// TIA Portal project "XSFW_TIA32801_A0" (V13) (continued)
REGION Network 3: Estado1-->Estado2 (Reposo--> Arranca cinta)
   RUNG wire#powerrail
      Contact( "1s1" )
      Contact( "iSNSpush_atras" )
      wire#w1
      Contact( "iS_automat" )
      wire#w2
      Contact( "iSNS_bs_abajo" )
      Contact( "Marcha" )
      wire#w3
      Contact( "Ya buscó caja" )
      wire#w4
      I_Contact( "Serie de Alarmas" )
      I_Contact( "Cajas acumuladas en salida" )
      Coil( "1c2" )
   END_RUNG
   RUNG wire#powerrail
      Contact( "1s8" )
      Contact( "CERO" )
      I_Contact( "Parada" )
      I_Contact( "Aux acaja acum" )
      I_Contact( "Aux caja trab" )
   END_RUNG wire#w1
   RUNG wire#w1
      Contact( "Modo Manual" )
      I_Contact( "iS_automat" )
      Contact( "fls_Modomanual" )
   END_RUNG wire#w2
   RUNG wire#w3
      Contact( "UNO" )
   END_RUNG wire#w4
   // the same network as SCL:
   "1c2" := (("1s1" AND "iSNSpush_atras") OR ("1s8" AND "CERO" AND NOT "Parada" AND NOT "Aux acaja acum" AND NOT "Aux caja trab")) AND ("iS_automat" OR ("Modo Manual" AND NOT "iS_automat" AND "fls_Modomanual")) AND "iSNS_bs_abajo" AND "Marcha" AND ("Ya buscó caja" OR "UNO") AND NOT "Serie de Alarmas" AND NOT "Cajas acumuladas en salida";
END_REGION

REGION Network 4: Estado2->Estado3 (Arranca Cinta --> Activar retenedores de caja)
   RUNG wire#powerrail
      { S7_Templates := "SrcType := DInt" } GE_Contact(in1 := "Encoder", in2 := 210)
      Contact( "1s2" )
      I_Contact( "Alarmas emergencia y térmicas" )
      I_Contact( "Alarmas cinta" )
      I_Contact( "Serie de Alarmas" )
      Coil( "1c3" )
   END_RUNG
   // the same network as SCL:
   "1c3" := ("Encoder" >= 210) AND "1s2" AND NOT "Alarmas emergencia y térmicas" AND NOT "Alarmas cinta" AND NOT "Serie de Alarmas";
END_REGION

REGION Network 5: Estado3-->Estado4 (Activar retenedores de caja--> Desactivar cinta)
   RUNG wire#powerrail
      Contact( "Punto neutro" )
      Contact( "1s3" )
      I_Contact( "Alarmas emergencia y térmicas" )
      I_Contact( "Alarmas cinta" )
      I_Contact( "Serie de Alarmas" )
      Coil( "1c4" )
   END_RUNG
   RUNG wire#powerrail
      { S7_Templates := "SrcType := DInt" } GE_Contact(in1 := "Encoder", in2 := 238)
      Coil( "Punto neutro" )
   END_RUNG
   // the same network as SCL:
   "1c4" := "Punto neutro" AND "1s3" AND NOT "Alarmas emergencia y térmicas" AND NOT "Alarmas cinta" AND NOT "Serie de Alarmas";
   "Punto neutro" := "Encoder" >= 238;
END_REGION

REGION Network 6: Estado4--> Estado5 (Desactivar cinta--> Activar Pusher y Pinza )
   RUNG wire#powerrail
      Contact( "1s4" )
      Contact( "Auxencol2" )
      I_Contact( "Alarmas"."falla en rele de cadena" )
      I_Contact( "Alarmas emergencia y térmicas" )
      I_Contact( "Alarmas salida y alim de cartones" )
      I_Contact( "Alarmas pusher" )
      I_Contact( "Alarmas brazo de succión" )
      I_Contact( "Serie de Alarmas" )
      Contact( "iSNSpush_atras" )
      Coil( "1c5" )
   END_RUNG
   // the same network as SCL:
   "1c5" := "1s4" AND "Auxencol2" AND NOT "Alarmas"."falla en rele de cadena" AND NOT "Alarmas emergencia y térmicas" AND NOT "Alarmas salida y alim de cartones" AND NOT "Alarmas pusher" AND NOT "Alarmas brazo de succión" AND NOT "Serie de Alarmas" AND "iSNSpush_atras";
END_REGION

REGION Network 7: Estado5-->Estado6 (Activar Pusher y Pinza--> Cilindro Pusher afuera)
   RUNG wire#powerrail
      Contact( "1s5" )
      wire#w1
      Contact( "iSNSalp" )
      I_Contact( "Serie de Alarmas" )
      I_Contact( "Alarmas emergencia y térmicas" )
      I_Contact( "Alarmas pusher" )
      Coil( "1c6" )
   END_RUNG
   RUNG wire#powerrail
      Contact( "CERO" )
      Contact( "1s3" )
      I_Contact( "1c4" )
   END_RUNG wire#w1
   RUNG wire#powerrail
      Contact( "CERO" )
      Contact( "1s4" )
      I_Contact( "1c5" )
   END_RUNG wire#w1
   // the same network as SCL:
   "1c6" := ("1s5" OR ("CERO" AND "1s3" AND NOT "1c4") OR ("CERO" AND "1s4" AND NOT "1c5")) AND "iSNSalp" AND NOT "Serie de Alarmas" AND NOT "Alarmas emergencia y térmicas" AND NOT "Alarmas pusher";
END_REGION

REGION Network 8: Estado6--> Estado7 (Cilindro Pusher afuera--> Desactivar cilindro pusher y pinza )
   RUNG wire#powerrail
      Contact( "1s6" )
      Contact( "iSNSpush_adel" )
      I_Contact( "Serie de Alarmas" )
      I_Contact( "Alarmas emergencia y térmicas" )
      I_Contact( "Alarmas pusher" )
      Coil( "1c7" )
   END_RUNG
   // the same network as SCL:
   "1c7" := "1s6" AND "iSNSpush_adel" AND NOT "Serie de Alarmas" AND NOT "Alarmas emergencia y térmicas" AND NOT "Alarmas pusher";
END_REGION

REGION Network 9: Estado7-->Estado8 (Desactivar cilindro pusher y pinza--> Área libre de Pusher)
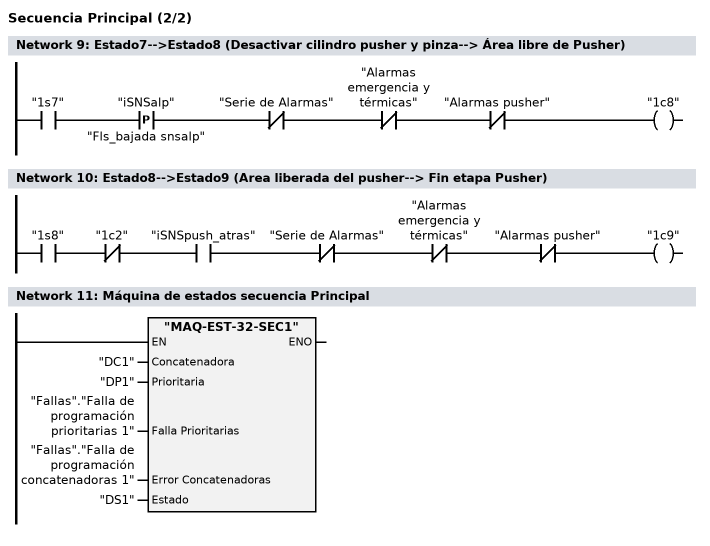
   RUNG wire#powerrail
      Contact( "1s7" )
      P_Contact(operand := "iSNSalp", bit := "Fls_bajada snsalp")
      I_Contact( "Serie de Alarmas" )
      I_Contact( "Alarmas emergencia y térmicas" )
      I_Contact( "Alarmas pusher" )
      Coil( "1c8" )
   END_RUNG
   // the same network as SCL:
   #_w1 := "1s7" AND "iSNSalp" AND NOT "Fls_bajada snsalp";   // rising edge of "iSNSalp"
   "Fls_bajada snsalp" := "iSNSalp";
   "1c8" := #_w1 AND NOT "Serie de Alarmas" AND NOT "Alarmas emergencia y térmicas" AND NOT "Alarmas pusher";
END_REGION

REGION Network 10: Estado8-->Estado9 (Area liberada del pusher--> Fin etapa Pusher)
   RUNG wire#powerrail
      Contact( "1s8" )
      I_Contact( "1c2" )
      Contact( "iSNSpush_atras" )
      I_Contact( "Serie de Alarmas" )
      I_Contact( "Alarmas emergencia y térmicas" )
      I_Contact( "Alarmas pusher" )
      Coil( "1c9" )
   END_RUNG
   // the same network as SCL:
   "1c9" := "1s8" AND NOT "1c2" AND "iSNSpush_atras" AND NOT "Serie de Alarmas" AND NOT "Alarmas emergencia y térmicas" AND NOT "Alarmas pusher";
END_REGION

REGION Network 11: Máquina de estados secuencia Principal
   RUNG wire#powerrail
      "MAQ-EST-32-SEC1"(Concatenadora := "DC1", Prioritaria := "DP1", "Falla Prioritarias" := "Fallas"."Falla de programación prioritarias 1", "Error Concatenadoras" := "Fallas"."Falla de programación concatenadoras 1", Estado := "DS1")
   END_RUNG
   // the same network as SCL:
   "MAQ-EST-32-SEC1"(Concatenadora := "DC1",
                     Prioritaria := "DP1",
                     "Falla Prioritarias" := "Fallas"."Falla de programación prioritarias 1",
                     "Error Concatenadoras" := "Fallas"."Falla de programación concatenadoras 1",
                     Estado := "DS1");
END_REGION
END_FUNCTION

FUNCTION "Condiciones de Marcha y Parada" : Void   // FC7, LAD
TITLE = Condiciones de MARCHA y PARADA (Se la considera una falla prioritaria).
{ S7_Optimized_Access := 'FALSE' }
VERSION : 0.1
// Establece la marcha del proceso según una determinada cantidad de condiciones. En particular para que arranque, se deberá presionar "avería/reposición" . Ya sea que se presione "Parada" o ocurra situaciones de Alarma, se desactivará "Marcha". La diferencia entre ambas es que, para arrancar el sistema luego de una parada, no hace falta presionar nuevamente "avería/reposición". Caso contrario ocurre si quiero arrancar el sistema luego de una Alarma.
BEGIN

REGION Network 1: Condiciones de Marcha
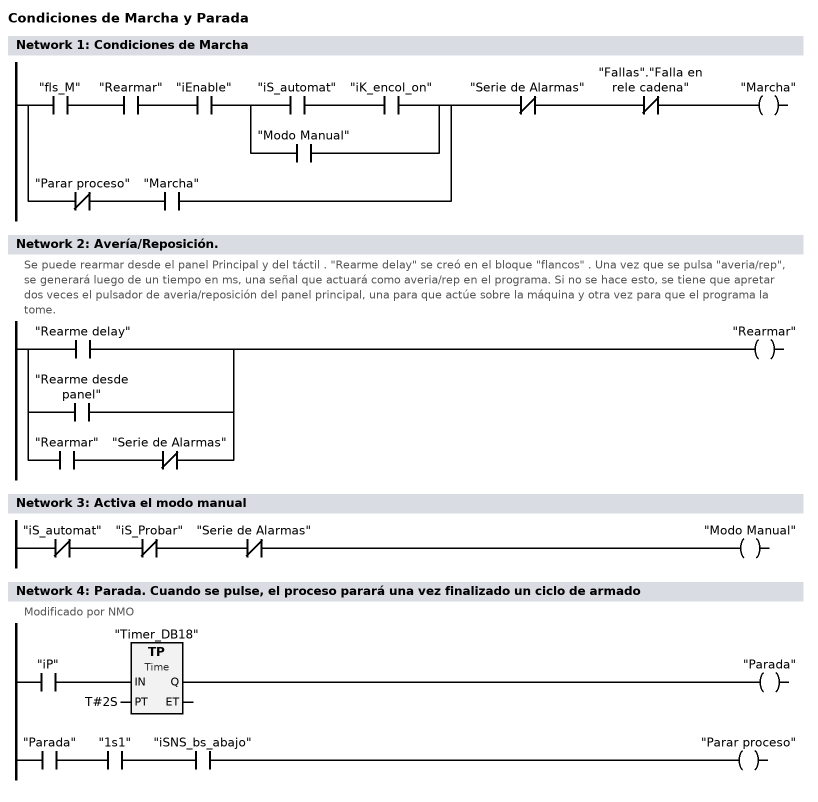
   RUNG wire#powerrail
      Contact( "fls_M" )
      Contact( "Rearmar" )
      Contact( "iEnable" )
      wire#w1
      Contact( "iS_automat" )
      Contact( "iK_encol_on" )
      wire#w2
      I_Contact( "Serie de Alarmas" )
      I_Contact( "Fallas"."Falla en rele cadena" )
      Coil( "Marcha" )
   END_RUNG
   RUNG wire#w1
      Contact( "Modo Manual" )
   END_RUNG wire#w2
   RUNG wire#powerrail
      I_Contact( "Parar proceso" )
      Contact( "Marcha" )
   END_RUNG wire#w2
   // the same network as SCL:
   "Marcha" := (("fls_M" AND "Rearmar" AND "iEnable" AND (("iS_automat" AND "iK_encol_on") OR "Modo Manual")) OR (NOT "Parar proceso" AND "Marcha")) AND NOT "Serie de Alarmas" AND NOT "Fallas"."Falla en rele cadena";
END_REGION

REGION Network 2: Avería/Reposición.
   // Se puede rearmar desde el panel Principal y del táctil . "Rearme delay" se creó en el bloque "flancos" . Una vez que se pulsa "averia/rep", se generará luego de un tiempo en ms, una señal que actuará como averia/rep en el programa. Si no se hace esto, se tiene que apretar dos veces el pulsador de averia/reposición del panel principal, una para que actúe sobre la máquina y otra vez para que el programa la tome.
   RUNG wire#powerrail
      Contact( "Rearme delay" )
      wire#w1
      Coil( "Rearmar" )
   END_RUNG
   RUNG wire#powerrail
      Contact( "Rearme desde panel" )
   END_RUNG wire#w1
   RUNG wire#powerrail
      Contact( "Rearmar" )
      I_Contact( "Serie de Alarmas" )
   END_RUNG wire#w1
   // the same network as SCL:
   "Rearmar" := "Rearme delay" OR "Rearme desde panel" OR ("Rearmar" AND NOT "Serie de Alarmas");
END_REGION

REGION Network 3: Activa el modo manual
   RUNG wire#powerrail
      I_Contact( "iS_automat" )
      I_Contact( "iS_Probar" )
      I_Contact( "Serie de Alarmas" )
      Coil( "Modo Manual" )
   END_RUNG
   // the same network as SCL:
   "Modo Manual" := NOT "iS_automat" AND NOT "iS_Probar" AND NOT "Serie de Alarmas";
END_REGION

REGION Network 4: Parada. Cuando se pulse, el proceso parará una vez finalizado un ciclo de armado
   // Modificado por NMO
   "Timer_DB18".TP(IN := "iP", PT := T#2S);
   "Parada" := "Timer_DB18".Q;
   "Parar proceso" := "Parada" AND "1s1" AND "iSNS_bs_abajo";
END_REGION
END_FUNCTION

FUNCTION "Contador rápido y encoder" : Void   // FC8, LAD
TITLE = Lleva la cuenta de los pulsos del ENCODER.
{ S7_Optimized_Access := 'FALSE' }
VERSION : 0.1
   VAR_TEMP   // added for the SCL form of the ladder/FBD networks
      _w1 : Bool;
   END_VAR
BEGIN

REGION Network 1: Reset del HSC para poner en cero el encóder.
   // En HSC va 258, es la ID de Hardware
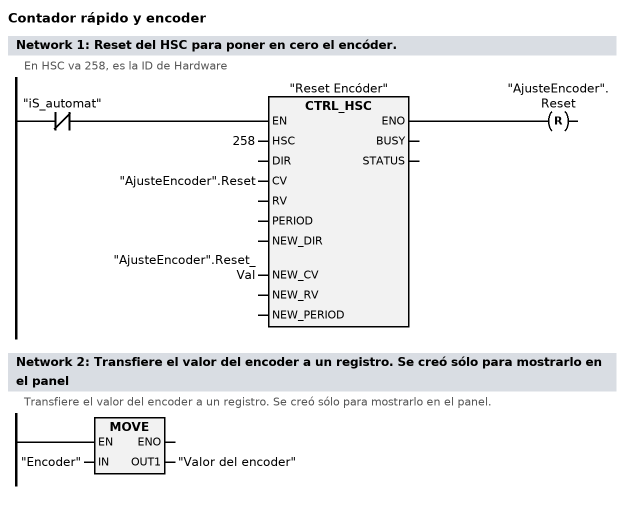
   // ENO of a box is taken as its EN; it also drops when the box reports an error
   #_w1 := NOT "iS_automat";
   IF #_w1 THEN
       "Reset Encóder"(HSC := 258, CV := "AjusteEncoder".Reset, NEW_CV := "AjusteEncoder".Reset_Val);   // CTRL_HSC
       "AjusteEncoder".Reset := FALSE;
   END_IF;
END_REGION

REGION Network 2: Transfiere el valor del encoder a un registro. Se creó sólo para mostrarlo en el panel
   // Transfiere el valor del encoder a un registro. Se creó sólo para mostrarlo en el panel.
   RUNG wire#powerrail
      { S7_GenerateENO := "TRUE" } Move(in := "Encoder", out1 => "Valor del encoder")
   END_RUNG
   // the same network as SCL:
   "Valor del encoder" := "Encoder";
END_REGION
END_FUNCTION

FUNCTION "cajas armadas hasta el momento" : Void   // FC9, LAD
{ S7_Optimized_Access := 'FALSE' }
VERSION : 0.1
BEGIN

REGION Network 1: Contabiliza la cantidad de cajas armadas.
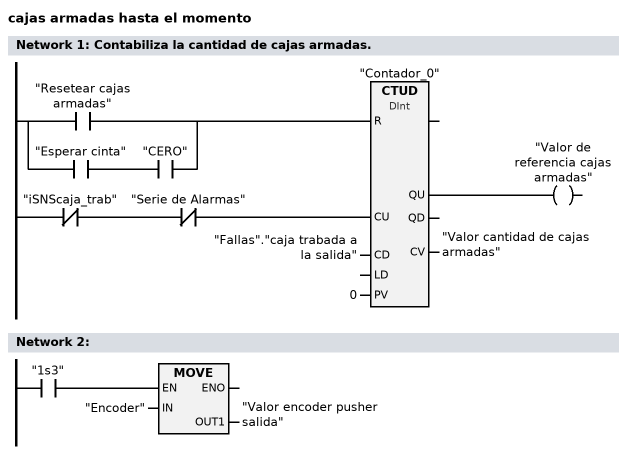
   "Contador_0".CTUD(cu := NOT "iSNScaja_trab" AND NOT "Serie de Alarmas",
                     r := "Resetear cajas armadas" OR ("Esperar cinta" AND "CERO"),
                     cd := "Fallas"."caja trabada a la salida",
                     pv := 0,
                     cv => "Valor cantidad de cajas armadas");
   "Valor de referencia cajas armadas" := "Contador_0".qu;
END_REGION

REGION Network 2
   RUNG wire#powerrail
      Contact( "1s3" )
      { S7_GenerateENO := "TRUE" } Move(in := "Encoder", out1 => "Valor encoder pusher salida")
   END_RUNG
   // the same network as SCL:
   IF "1s3" THEN "Valor encoder pusher salida" := "Encoder"; END_IF;
END_REGION
END_FUNCTION

FUNCTION "Luces de marcha y parada" : Void   // FC10, LAD
{ S7_Optimized_Access := 'FALSE' }
VERSION : 0.1
BEGIN

REGION Network 1: Luz de Marcha
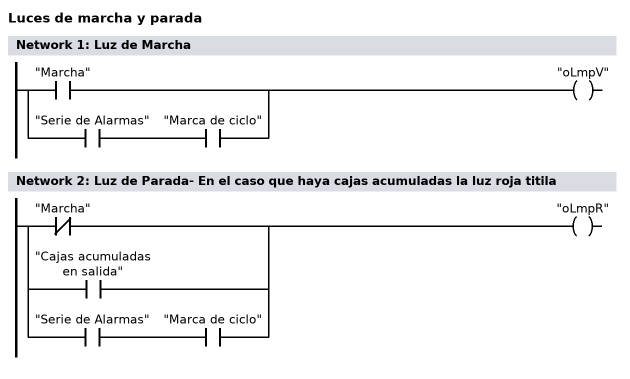
   RUNG wire#powerrail
      Contact( "Marcha" )
      wire#w1
      Coil( "oLmpV" )
   END_RUNG
   RUNG wire#powerrail
      Contact( "Serie de Alarmas" )
      Contact( "Marca de ciclo" )
   END_RUNG wire#w1
   // the same network as SCL:
   "oLmpV" := "Marcha" OR ("Serie de Alarmas" AND "Marca de ciclo");
END_REGION

REGION Network 2: Luz de Parada- En el caso que haya cajas acumuladas la luz roja titila
   RUNG wire#powerrail
      I_Contact( "Marcha" )
      wire#w1
      Coil( "oLmpR" )
   END_RUNG
   RUNG wire#powerrail
      Contact( "Cajas acumuladas en salida" )
   END_RUNG wire#w1
   RUNG wire#powerrail
      Contact( "Serie de Alarmas" )
      Contact( "Marca de ciclo" )
   END_RUNG wire#w1
   // the same network as SCL:
   "oLmpR" := NOT "Marcha" OR "Cajas acumuladas en salida" OR ("Serie de Alarmas" AND "Marca de ciclo");
END_REGION
END_FUNCTION

FUNCTION "flancos" : Void   // FC12, LAD
{ S7_Optimized_Access := 'FALSE' }
VERSION : 0.1
   VAR_TEMP   // added for the SCL form of the ladder/FBD networks
      _w1 : Bool;
   END_VAR
BEGIN

REGION Network 1: avería/ reposición
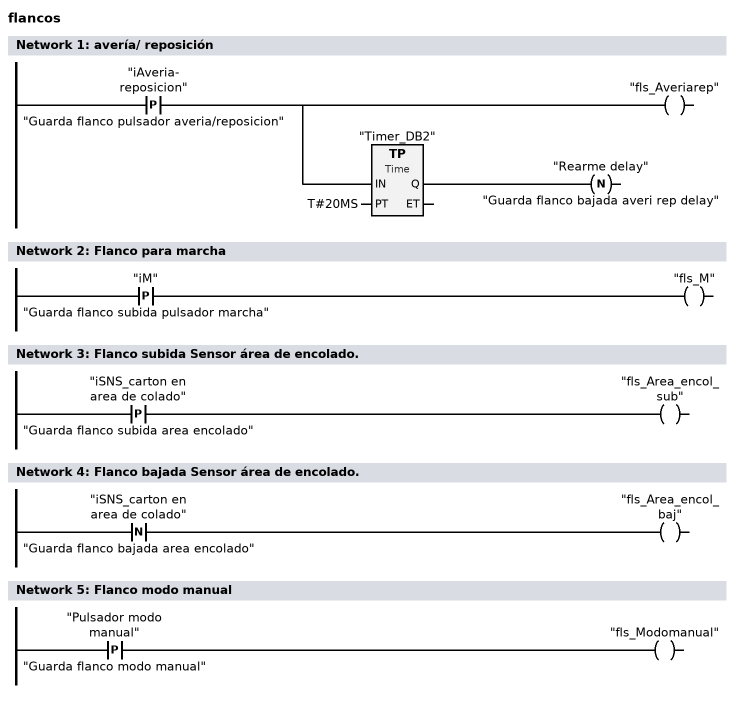
   #_w1 := "iAveria-reposicion" AND NOT "Guarda flanco pulsador averia/reposicion";   // rising edge of "iAveria-reposicion"
   "Guarda flanco pulsador averia/reposicion" := "iAveria-reposicion";
   "fls_Averiarep" := #_w1;
   "Timer_DB2".TP(in := #_w1, pt := T#20MS);
   "Rearme delay" := NOT "Timer_DB2".q AND "Guarda flanco bajada averi rep delay";   // falling edge
   "Guarda flanco bajada averi rep delay" := "Timer_DB2".q;
END_REGION

REGION Network 2: Flanco para marcha
   RUNG wire#powerrail
      P_Contact(operand := "iM", bit := "Guarda flanco subida pulsador marcha")
      Coil( "fls_M" )
   END_RUNG
   // the same network as SCL:
   #_w1 := "iM" AND NOT "Guarda flanco subida pulsador marcha";   // rising edge of "iM"
   "Guarda flanco subida pulsador marcha" := "iM";
   "fls_M" := #_w1;
END_REGION

REGION Network 3: Flanco subida Sensor área de encolado.
   RUNG wire#powerrail
      P_Contact(operand := "iSNS_carton en area de colado", bit := "Guarda flanco subida area encolado")
      Coil( "fls_Area_encol_sub" )
   END_RUNG
   // the same network as SCL:
   #_w1 := "iSNS_carton en area de colado" AND NOT "Guarda flanco subida area encolado";   // rising edge of "iSNS_carton en area de colado"
   "Guarda flanco subida area encolado" := "iSNS_carton en area de colado";
   "fls_Area_encol_sub" := #_w1;
END_REGION

REGION Network 4: Flanco bajada Sensor área de encolado.
   RUNG wire#powerrail
      N_Contact(operand := "iSNS_carton en area de colado", bit := "Guarda flanco bajada area encolado")
      Coil( "fls_Area_encol_baj" )
   END_RUNG
   // the same network as SCL:
   #_w1 := NOT "iSNS_carton en area de colado" AND "Guarda flanco bajada area encolado";   // falling edge of "iSNS_carton en area de colado"
   "Guarda flanco bajada area encolado" := "iSNS_carton en area de colado";
   "fls_Area_encol_baj" := #_w1;
END_REGION

REGION Network 5: Flanco modo manual
   RUNG wire#powerrail
      P_Contact(operand := "Pulsador modo manual", bit := "Guarda flanco modo manual")
      Coil( "fls_Modomanual" )
   END_RUNG
   // the same network as SCL:
   #_w1 := "Pulsador modo manual" AND NOT "Guarda flanco modo manual";   // rising edge of "Pulsador modo manual"
   "Guarda flanco modo manual" := "Pulsador modo manual";
   "fls_Modomanual" := #_w1;
END_REGION
END_FUNCTION

FUNCTION "MODO PROBAR (MP)" : Void   // FC13, LAD
{ S7_Optimized_Access := 'FALSE' }
VERSION : 0.1
   VAR_TEMP   // added for the SCL form of the ladder/FBD networks
      _w1 : Bool;
   END_VAR
BEGIN

REGION Network 1: Modo Probar. En este caso se desactivan las alarmas excepto la de emergencia y térmicas.
   // Si no está en automático, y no hay alarmas, se activa el modo PROBAR. Con esto se activa la bomba de vacío.
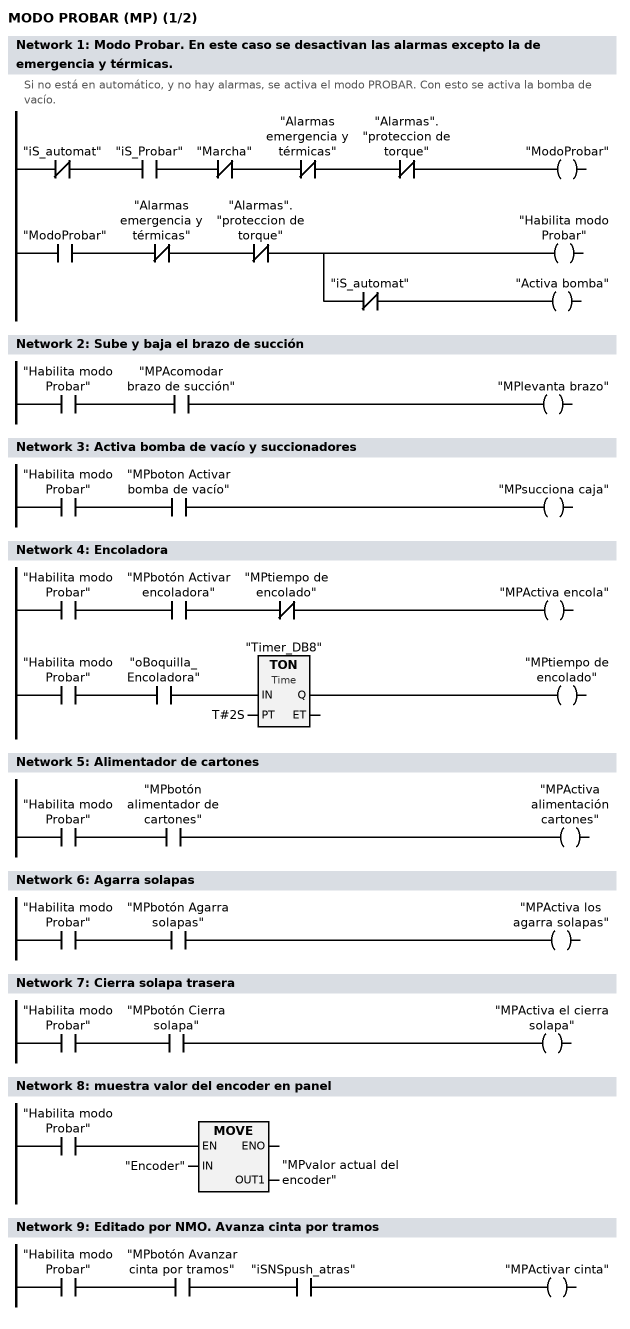
   RUNG wire#powerrail
      I_Contact( "iS_automat" )
      Contact( "iS_Probar" )
      I_Contact( "Marcha" )
      I_Contact( "Alarmas emergencia y térmicas" )
      I_Contact( "Alarmas"."proteccion de torque" )
      Coil( "ModoProbar" )
   END_RUNG
   RUNG wire#powerrail
      Contact( "ModoProbar" )
      I_Contact( "Alarmas emergencia y térmicas" )
      I_Contact( "Alarmas"."proteccion de torque" )
      wire#w1
      Coil( "Habilita modo Probar" )
   END_RUNG
   RUNG wire#w1
      I_Contact( "iS_automat" )
      Coil( "Activa bomba" )
   END_RUNG
   // the same network as SCL:
   "ModoProbar" := NOT "iS_automat" AND "iS_Probar" AND NOT "Marcha" AND NOT "Alarmas emergencia y térmicas" AND NOT "Alarmas"."proteccion de torque";
   "Habilita modo Probar" := "ModoProbar" AND NOT "Alarmas emergencia y térmicas" AND NOT "Alarmas"."proteccion de torque";
   "Activa bomba" := "Habilita modo Probar" AND NOT "iS_automat";
END_REGION

REGION Network 2: Sube y baja el brazo de succión
   RUNG wire#powerrail
      Contact( "Habilita modo Probar" )
      Contact( "MPAcomodar brazo de succión" )
      Coil( "MPlevanta brazo" )
   END_RUNG
   // the same network as SCL:
   "MPlevanta brazo" := "Habilita modo Probar" AND "MPAcomodar brazo de succión";
END_REGION

REGION Network 3: Activa bomba de vacío y succionadores
   RUNG wire#powerrail
      Contact( "Habilita modo Probar" )
      Contact( "MPboton Activar bomba de vacío" )
      Coil( "MPsucciona caja" )
   END_RUNG
   // the same network as SCL:
   "MPsucciona caja" := "Habilita modo Probar" AND "MPboton Activar bomba de vacío";
END_REGION

REGION Network 4: Encoladora
   "MPActiva encola" := "Habilita modo Probar" AND "MPbotón Activar encoladora" AND NOT "MPtiempo de encolado";
   "Timer_DB8".TON(IN := "Habilita modo Probar" AND "oBoquilla_Encoladora", PT := T#2S);
   "MPtiempo de encolado" := "Timer_DB8".Q;
END_REGION

REGION Network 5: Alimentador de cartones
   RUNG wire#powerrail
      Contact( "Habilita modo Probar" )
      Contact( "MPbotón alimentador de cartones" )
      Coil( "MPActiva alimentación cartones" )
   END_RUNG
   // the same network as SCL:
   "MPActiva alimentación cartones" := "Habilita modo Probar" AND "MPbotón alimentador de cartones";
END_REGION

REGION Network 6: Agarra solapas
   RUNG wire#powerrail
      Contact( "Habilita modo Probar" )
      Contact( "MPbotón Agarra solapas" )
      Coil( "MPActiva los agarra solapas" )
   END_RUNG
   // the same network as SCL:
   "MPActiva los agarra solapas" := "Habilita modo Probar" AND "MPbotón Agarra solapas";
END_REGION

REGION Network 7: Cierra solapa trasera
   RUNG wire#powerrail
      Contact( "Habilita modo Probar" )
      Contact( "MPbotón Cierra solapa" )
      Coil( "MPActiva el cierra solapa" )
   END_RUNG
   // the same network as SCL:
   "MPActiva el cierra solapa" := "Habilita modo Probar" AND "MPbotón Cierra solapa";
END_REGION

REGION Network 8: muestra valor del encoder en panel
   RUNG wire#powerrail
      Contact( "Habilita modo Probar" )
      { S7_GenerateENO := "TRUE" } Move(in := "Encoder", out1 => "MPvalor actual del encoder")
   END_RUNG
   // the same network as SCL:
   IF "Habilita modo Probar" THEN "MPvalor actual del encoder" := "Encoder"; END_IF;
END_REGION

REGION Network 9: Editado por NMO. Avanza cinta por tramos
   RUNG wire#powerrail
      Contact( "Habilita modo Probar" )
      Contact( "MPbotón Avanzar cinta por tramos" )
      Contact( "iSNSpush_atras" )
      Coil( "MPActivar cinta" )
   END_RUNG
   // the same network as SCL:
   "MPActivar cinta" := "Habilita modo Probar" AND "MPbotón Avanzar cinta por tramos" AND "iSNSpush_atras";
END_REGION

REGION Network 10: Editado por NMO. Desactivar marca "MPbotón avanzar cinta por tramos".
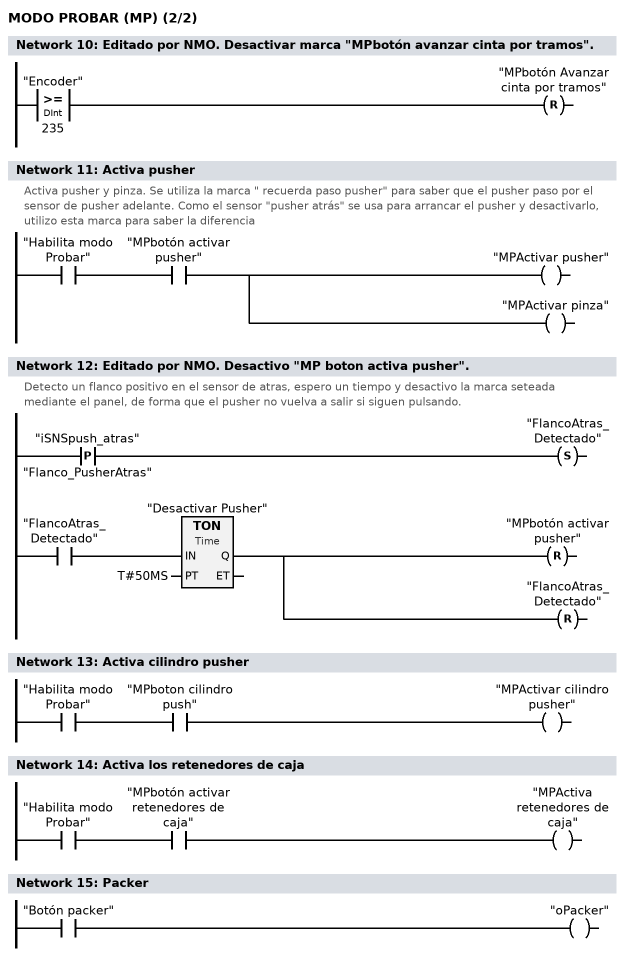
   RUNG wire#powerrail
      { S7_Templates := "SrcType := DInt" } GE_Contact(in1 := "Encoder", in2 := 235)
      R_Coil( "MPbotón Avanzar cinta por tramos" )
   END_RUNG
   // the same network as SCL:
   IF "Encoder" >= 235 THEN "MPbotón Avanzar cinta por tramos" := FALSE; END_IF;
END_REGION

REGION Network 11: Activa pusher
   // Activa pusher y pinza. Se utiliza la marca " recuerda paso pusher" para saber que el pusher paso por el sensor de pusher adelante. Como el sensor "pusher atrás" se usa para arrancar el pusher y desactivarlo, utilizo esta marca para saber la diferencia
   RUNG wire#powerrail
      Contact( "Habilita modo Probar" )
      Contact( "MPbotón activar pusher" )
      wire#w1
      Coil( "MPActivar pusher" )
   END_RUNG
   RUNG wire#w1
      Coil( "MPActivar pinza" )
   END_RUNG
   // the same network as SCL:
   "MPActivar pusher" := "Habilita modo Probar" AND "MPbotón activar pusher";
   "MPActivar pinza" := "MPActivar pusher";
END_REGION

REGION Network 12: Editado por NMO. Desactivo "MP boton activa pusher".
   // Detecto un flanco positivo en el sensor de atras, espero un tiempo y desactivo la marca seteada mediante el panel, de forma que el pusher no vuelva a salir si siguen pulsando.
   #_w1 := "iSNSpush_atras" AND NOT "Flanco_PusherAtras";   // rising edge of "iSNSpush_atras"
   "Flanco_PusherAtras" := "iSNSpush_atras";
   IF #_w1 THEN "FlancoAtras_Detectado" := TRUE; END_IF;
   "Desactivar Pusher".TON(IN := "FlancoAtras_Detectado", PT := T#50MS);
   IF "Desactivar Pusher".Q THEN
       "MPbotón activar pusher" := FALSE;
       "FlancoAtras_Detectado" := FALSE;
   END_IF;
END_REGION

REGION Network 13: Activa cilindro pusher
   RUNG wire#powerrail
      Contact( "Habilita modo Probar" )
      Contact( "MPboton cilindro push" )
      Coil( "MPActivar cilindro pusher" )
   END_RUNG
   // the same network as SCL:
   "MPActivar cilindro pusher" := "Habilita modo Probar" AND "MPboton cilindro push";
END_REGION

REGION Network 14: Activa los retenedores de caja
   RUNG wire#powerrail
      Contact( "Habilita modo Probar" )
      Contact( "MPbotón activar retenedores de caja" )
      Coil( "MPActiva retenedores de caja" )
   END_RUNG
   // the same network as SCL:
   "MPActiva retenedores de caja" := "Habilita modo Probar" AND "MPbotón activar retenedores de caja";
END_REGION

REGION Network 15: Packer
   RUNG wire#powerrail
      Contact( "Botón packer" )
      Coil( "oPacker" )
   END_RUNG
   // the same network as SCL:
   "oPacker" := "Botón packer";
END_REGION
END_FUNCTION

FUNCTION "Tratamiento de Fallas" : Void   // FC16, LAD
TITLE = Tratamiento de fallas.
{ S7_Optimized_Access := 'FALSE' }
VERSION : 0.1
   VAR_TEMP   // added for the SCL form of the ladder/FBD networks
      _w1 : Bool;
   END_VAR
BEGIN

REGION Network 1: Falla en térmicas.
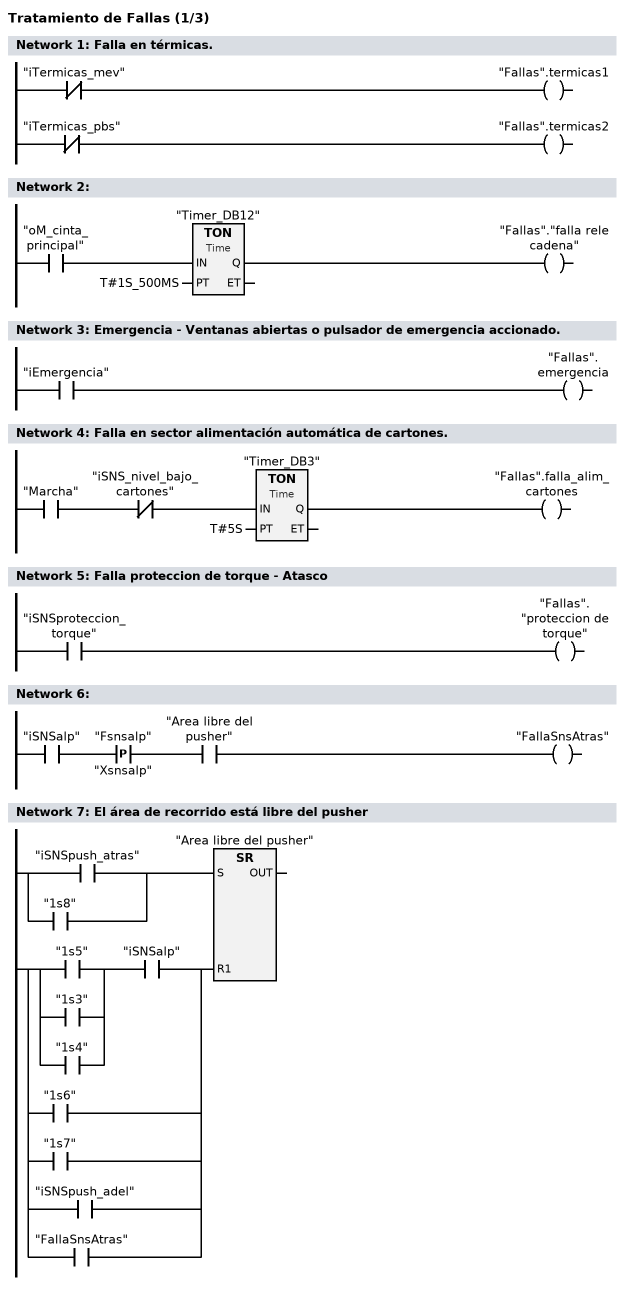
   RUNG wire#powerrail
      I_Contact( "iTermicas_mev" )
      Coil( "Fallas".termicas1 )
   END_RUNG
   RUNG wire#powerrail
      I_Contact( "iTermicas_pbs" )
      Coil( "Fallas".termicas2 )
   END_RUNG
   // the same network as SCL:
   "Fallas".termicas1 := NOT "iTermicas_mev";
   "Fallas".termicas2 := NOT "iTermicas_pbs";
END_REGION

REGION Network 2
   "Timer_DB12".TON(IN := "oM_cinta_principal", PT := T#1S_500MS);
   "Fallas"."falla rele cadena" := "Timer_DB12".Q;
END_REGION

REGION Network 3: Emergencia - Ventanas abiertas o pulsador de emergencia accionado.
   RUNG wire#powerrail
      Contact( "iEmergencia" )
      Coil( "Fallas".emergencia )
   END_RUNG
   // the same network as SCL:
   "Fallas".emergencia := "iEmergencia";
END_REGION

REGION Network 4: Falla en sector alimentación automática de cartones.
   "Timer_DB3".TON(IN := "Marcha" AND NOT "iSNS_nivel_bajo_cartones", PT := T#5S);
   "Fallas".falla_alim_cartones := "Timer_DB3".Q;
END_REGION

REGION Network 5: Falla proteccion de torque - Atasco
   RUNG wire#powerrail
      Contact( "iSNSproteccion_torque" )
      Coil( "Fallas"."proteccion de torque" )
   END_RUNG
   // the same network as SCL:
   "Fallas"."proteccion de torque" := "iSNSproteccion_torque";
END_REGION

REGION Network 6
   RUNG wire#powerrail
      Contact( "iSNSalp" )
      P_Contact(operand := "Fsnsalp", bit := "Xsnsalp")
      Contact( "Area libre del pusher" )
      Coil( "FallaSnsAtras" )
   END_RUNG
   // the same network as SCL:
   #_w1 := "iSNSalp" AND "Fsnsalp" AND NOT "Xsnsalp";   // rising edge of "Fsnsalp"
   "Xsnsalp" := "Fsnsalp";
   "FallaSnsAtras" := #_w1 AND "Area libre del pusher";
END_REGION

REGION Network 7: El área de recorrido está libre del pusher
   RUNG wire#powerrail
      Contact( "iSNSpush_atras" )
      wire#w1
      S_SR(operand := "Area libre del pusher", r1 := wire#w3)
   END_RUNG
   RUNG wire#powerrail
      Contact( "1s8" )
   END_RUNG wire#w1
   RUNG wire#powerrail
      Contact( "1s5" )
      wire#w2
      Contact( "iSNSalp" )
   END_RUNG wire#w3
   RUNG wire#powerrail
      Contact( "1s3" )
   END_RUNG wire#w2
   RUNG wire#powerrail
      Contact( "1s4" )
   END_RUNG wire#w2
   RUNG wire#powerrail
      Contact( "1s6" )
   END_RUNG wire#w3
   RUNG wire#powerrail
      Contact( "1s7" )
   END_RUNG wire#w3
   RUNG wire#powerrail
      Contact( "iSNSpush_adel" )
   END_RUNG wire#w3
   RUNG wire#powerrail
      Contact( "FallaSnsAtras" )
   END_RUNG wire#w3
   // the same network as SCL:
   IF "iSNSpush_atras" OR "1s8" THEN
       "Area libre del pusher" := TRUE;   // SR flip-flop
   END_IF;
   IF (("1s5" OR "1s3" OR "1s4") AND "iSNSalp") OR "1s6" OR "1s7" OR "iSNSpush_adel" OR "FallaSnsAtras" THEN
       "Area libre del pusher" := FALSE;
   END_IF;
END_REGION

REGION Network 8: Incongruencia en sensores del pusher.
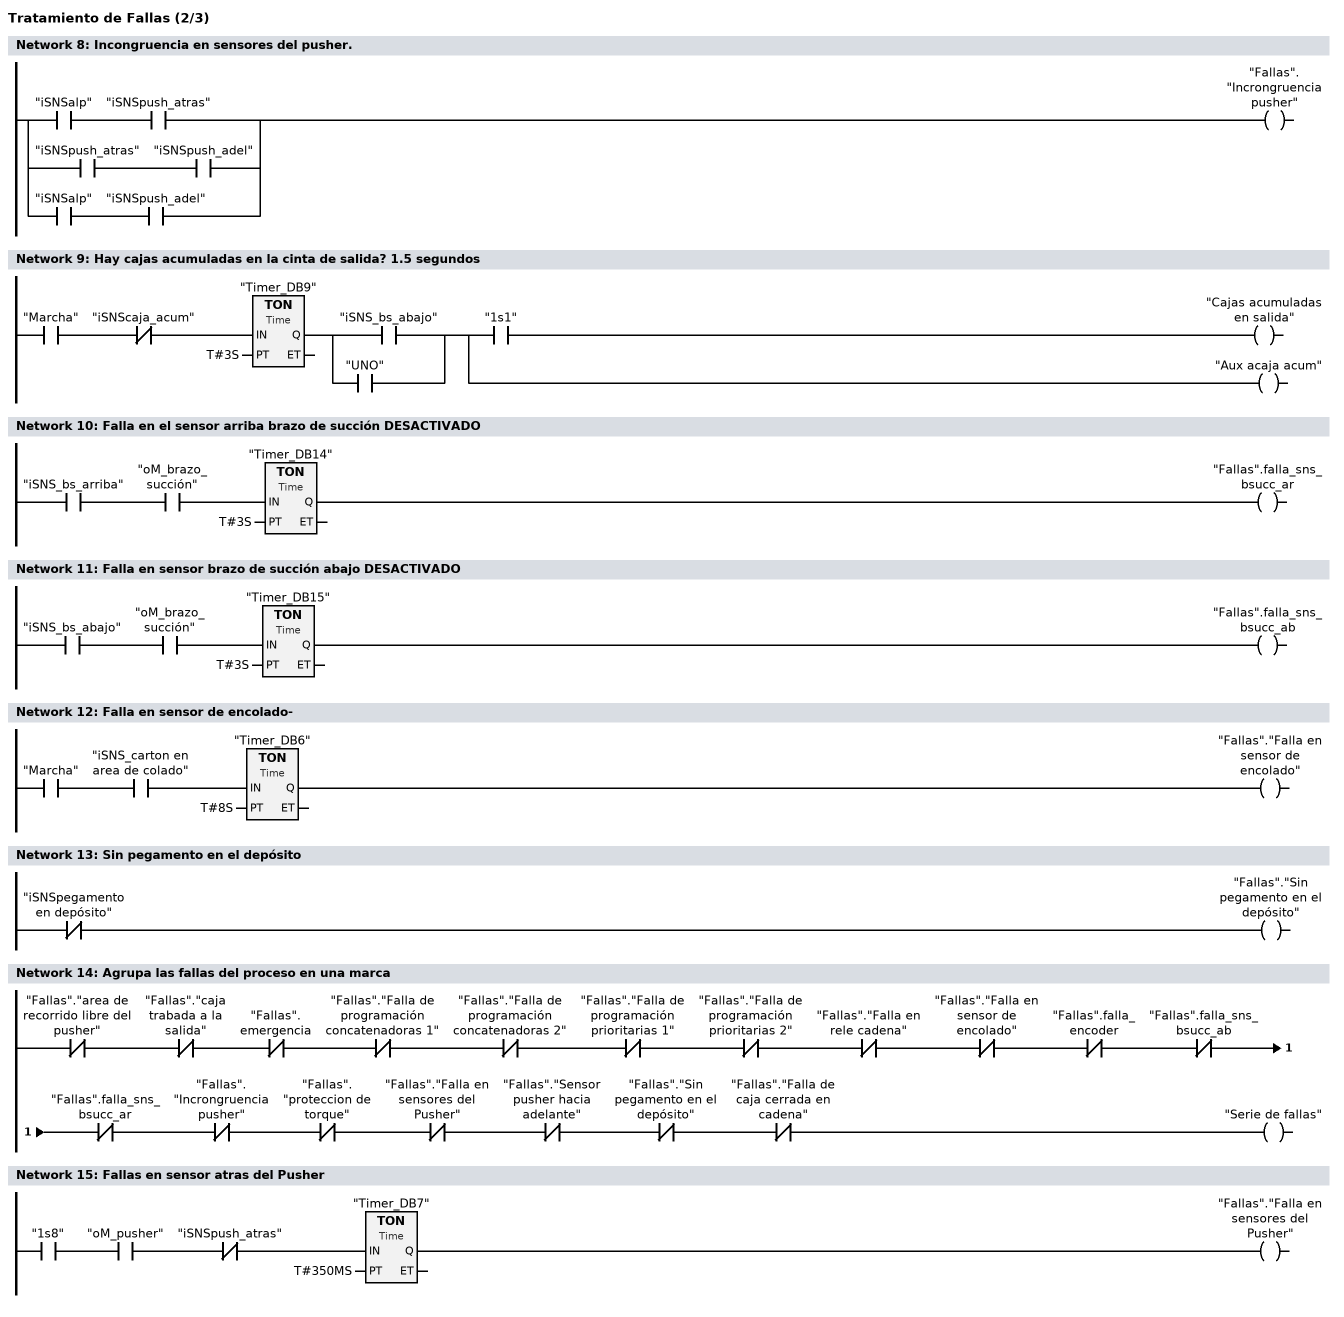
   RUNG wire#powerrail
      Contact( "iSNSalp" )
      Contact( "iSNSpush_atras" )
      wire#w1
      Coil( "Fallas"."Incrongruencia pusher" )
   END_RUNG
   RUNG wire#powerrail
      Contact( "iSNSpush_atras" )
      Contact( "iSNSpush_adel" )
   END_RUNG wire#w1
   RUNG wire#powerrail
      Contact( "iSNSalp" )
      Contact( "iSNSpush_adel" )
   END_RUNG wire#w1
   // the same network as SCL:
   "Fallas"."Incrongruencia pusher" := ("iSNSalp" AND "iSNSpush_atras") OR ("iSNSpush_atras" AND "iSNSpush_adel") OR ("iSNSalp" AND "iSNSpush_adel");
END_REGION

REGION Network 9: Hay cajas acumuladas en la cinta de salida? 1.5 segundos
   "Timer_DB9".TON(in := "Marcha" AND NOT "iSNScaja_acum", pt := T#3S);
   #_w1 := "Timer_DB9".q AND ("iSNS_bs_abajo" OR "UNO");
   "Cajas acumuladas en salida" := #_w1 AND "1s1";
   "Aux acaja acum" := #_w1;
END_REGION

REGION Network 10: Falla en el sensor arriba brazo de succión DESACTIVADO
   "Timer_DB14".TON(IN := "iSNS_bs_arriba" AND "oM_brazo_succión", PT := T#3S);
   "Fallas".falla_sns_bsucc_ar := "Timer_DB14".Q;
END_REGION

REGION Network 11: Falla en sensor brazo de succión abajo DESACTIVADO
   "Timer_DB15".TON(IN := "iSNS_bs_abajo" AND "oM_brazo_succión", PT := T#3S);
   "Fallas".falla_sns_bsucc_ab := "Timer_DB15".Q;
END_REGION

REGION Network 12: Falla en sensor de encolado-
   "Timer_DB6".TON(IN := "Marcha" AND "iSNS_carton en area de colado", PT := T#8S);
   "Fallas"."Falla en sensor de encolado" := "Timer_DB6".Q;
END_REGION

REGION Network 13: Sin pegamento en el depósito
   RUNG wire#powerrail
      I_Contact( "iSNSpegamento en depósito" )
      Coil( "Fallas"."Sin pegamento en el depósito" )
   END_RUNG
   // the same network as SCL:
   "Fallas"."Sin pegamento en el depósito" := NOT "iSNSpegamento en depósito";
END_REGION

REGION Network 14: Agrupa las fallas del proceso en una marca
   RUNG wire#powerrail
      I_Contact( "Fallas"."area de recorrido libre del pusher" )
      I_Contact( "Fallas"."caja trabada a la salida" )
      I_Contact( "Fallas".emergencia )
      I_Contact( "Fallas"."Falla de programación concatenadoras 1" )
      I_Contact( "Fallas"."Falla de programación concatenadoras 2" )
      I_Contact( "Fallas"."Falla de programación prioritarias 1" )
      I_Contact( "Fallas"."Falla de programación prioritarias 2" )
      I_Contact( "Fallas"."Falla en rele cadena" )
      I_Contact( "Fallas"."Falla en sensor de encolado" )
      I_Contact( "Fallas".falla_encoder )
      I_Contact( "Fallas".falla_sns_bsucc_ab )
      I_Contact( "Fallas".falla_sns_bsucc_ar )
      I_Contact( "Fallas"."Incrongruencia pusher" )
      I_Contact( "Fallas"."proteccion de torque" )
      I_Contact( "Fallas"."Falla en sensores del Pusher" )
      I_Contact( "Fallas"."Sensor pusher hacia adelante" )
      I_Contact( "Fallas"."Sin pegamento en el depósito" )
      I_Contact( "Fallas"."Falla de caja cerrada en cadena" )
      Coil( "Serie de fallas" )
   END_RUNG
   // the same network as SCL:
   "Serie de fallas" := NOT "Fallas"."area de recorrido libre del pusher" AND NOT "Fallas"."caja trabada a la salida" AND NOT "Fallas".emergencia AND NOT "Fallas"."Falla de programación concatenadoras 1" AND NOT "Fallas"."Falla de programación concatenadoras 2" AND NOT "Fallas"."Falla de programación prioritarias 1" AND NOT "Fallas"."Falla de programación prioritarias 2" AND NOT "Fallas"."Falla en rele cadena" AND NOT "Fallas"."Falla en sensor de encolado" AND NOT "Fallas".falla_encoder AND NOT "Fallas".falla_sns_bsucc_ab AND NOT "Fallas".falla_sns_bsucc_ar AND NOT "Fallas"."Incrongruencia pusher" AND NOT "Fallas"."proteccion de torque" AND NOT "Fallas"."Falla en sensores del Pusher" AND NOT "Fallas"."Sensor pusher hacia adelante" AND NOT "Fallas"."Sin pegamento en el depósito" AND NOT "Fallas"."Falla de caja cerrada en cadena";
END_REGION

REGION Network 15: Fallas en sensor atras del Pusher
   "Timer_DB7".TON(IN := "1s8" AND "oM_pusher" AND NOT "iSNSpush_atras", PT := T#350MS);
   "Fallas"."Falla en sensores del Pusher" := "Timer_DB7".Q;
END_REGION

REGION Network 16: Fallas en sensor adelante del Pusher
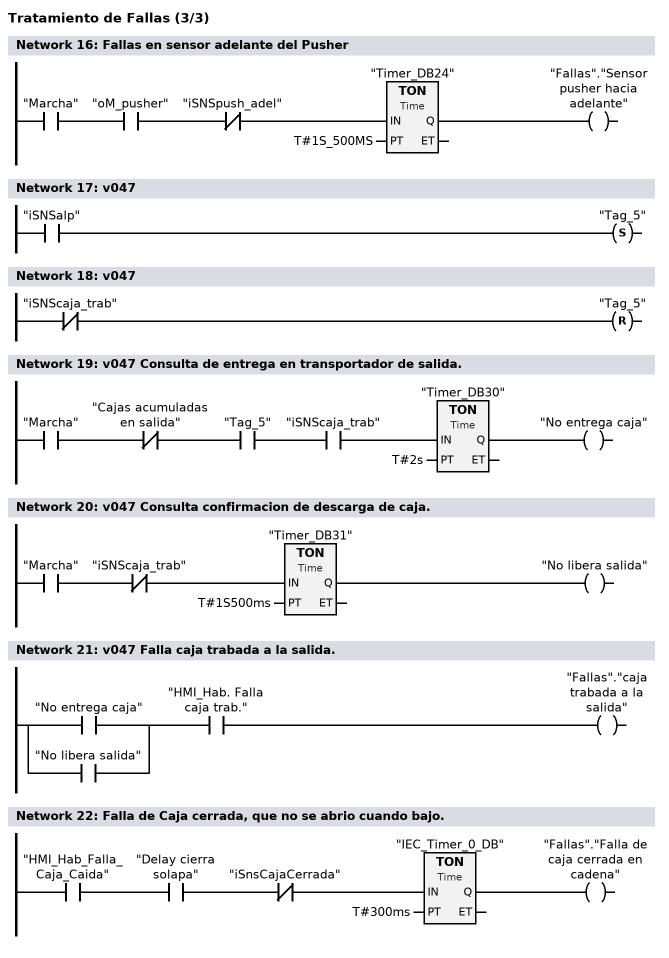
   "Timer_DB24".TON(IN := "Marcha" AND "oM_pusher" AND NOT "iSNSpush_adel", PT := T#1S_500MS);
   "Fallas"."Sensor pusher hacia adelante" := "Timer_DB24".Q;
END_REGION

REGION Network 17: v047
   RUNG wire#powerrail
      Contact( "iSNSalp" )
      S_Coil( "Tag_5" )
   END_RUNG
   // the same network as SCL:
   IF "iSNSalp" THEN "Tag_5" := TRUE; END_IF;
END_REGION

REGION Network 18: v047
   RUNG wire#powerrail
      I_Contact( "iSNScaja_trab" )
      R_Coil( "Tag_5" )
   END_RUNG
   // the same network as SCL:
   IF NOT "iSNScaja_trab" THEN "Tag_5" := FALSE; END_IF;
END_REGION

REGION Network 19: v047 Consulta de entrega en transportador de salida.
   "Timer_DB30".TON(IN := "Marcha" AND NOT "Cajas acumuladas en salida" AND "Tag_5" AND "iSNScaja_trab",
                    PT := T#2s);
   "No entrega caja" := "Timer_DB30".Q;
END_REGION

REGION Network 20: v047 Consulta confirmacion de descarga de caja.
   "Timer_DB31".TON(IN := "Marcha" AND NOT "iSNScaja_trab", PT := T#1S500ms);
   "No libera salida" := "Timer_DB31".Q;
END_REGION

REGION Network 21: v047 Falla caja trabada a la salida.
   RUNG wire#powerrail
      Contact( "No entrega caja" )
      wire#w1
      Contact( "HMI_Hab. Falla caja trab." )
      Coil( "Fallas"."caja trabada a la salida" )
   END_RUNG
   RUNG wire#powerrail
      Contact( "No libera salida" )
   END_RUNG wire#w1
   // the same network as SCL:
   "Fallas"."caja trabada a la salida" := ("No entrega caja" OR "No libera salida") AND "HMI_Hab. Falla caja trab.";
END_REGION

REGION Network 22: Falla de Caja cerrada, que no se abrio cuando bajo.
   "IEC_Timer_0_DB".TON(IN := "HMI_Hab_Falla_Caja_Caida" AND "Delay cierra solapa" AND NOT "iSnsCajaCerrada",
                        PT := T#300ms);
   "Fallas"."Falla de caja cerrada en cadena" := "IEC_Timer_0_DB".Q;
END_REGION
END_FUNCTION

FUNCTION "Salidas" : Void   // FC17, LAD
TITLE = Salidas del proceso (Modo Automático y Manual)
{ S7_Optimized_Access := 'FALSE' }
VERSION : 0.1
   VAR_TEMP   // added for the SCL form of the ladder/FBD networks
      _w1 : Bool;
   END_VAR
BEGIN

REGION Network 1: Activa la línea de emergencia del PLC